   12103: 'Pump1: FeedPump: max. filling level drip pan', class Pump Warning Alarm, trigger "Pump1_FeedPump_DBW_2" bit 10
   12104: 'Pump1: FeedPump: dry-run protection', class Pump Warning Alarm, trigger "Pump1_FeedPump_DBW_2" bit 11
   12105: 'Pump1: FeedPump: incorrect time entry for runtime or pause time', class Pump Warning Alarm, trigger "Pump1_FeedPump_DBW_2" bit 12
   12106: 'Pump1: FeedPump: temperature for switch-off not reached', class Pump Warning Alarm, trigger "Pump1_FeedPump_DBW_2" bit 13
   12107: 'Pump1: FeedPump: fan motor protecting switch', class Pump Warning Alarm, trigger "Pump1_FeedPump_DBW_2" bit 14
   12108: 'Pump1: FeedPump: filling level too low', class Pump Warning Alarm, trigger "Pump1_FeedPump_DBW_2" bit 15
   12109: 'Pump1: FeedPump:', class Pump Warning Alarm, trigger "Pump1_FeedPump_DBW_2" bit 0
   12110: 'Pump1: FeedPump: filling selected but no barrel present', class Pump Warning Alarm, trigger "Pump1_FeedPump_DBW_2" bit 1
   12111: 'Pump1: FeedPump: no barrel present', class Pump Warning Alarm, trigger "Pump1_FeedPump_DBW_2" bit 2
   12112: 'Pump1: FeedPump:', class Pump Warning Alarm, trigger "Pump1_EdgeFilter_DBW_28" bit 8
   12113: 'Pump1: EdgeFilter: motor protecting switch has tripped', class Pump Warning Alarm, trigger "Pump1_EdgeFilter_DBW_28" bit 9
   12114: 'Pump1: EdgeFilter: max. differential pressure', class Pump Warning Alarm, trigger "Pump1_EdgeFilter_DBW_28" bit 10
   12115: 'Pump1: EdgeFilter: incorrect time entry for runtime or pause time', class Pump Warning Alarm, trigger "Pump1_EdgeFilter_DBW_28" bit 11
   12117: 'Pump1: Component pump: admission pressure not present', class Pump Archive Error Foaming, trigger "Pump1_Component_DBW_56" bit 8
   12118: 'Pump1: Component pump: motor protecting switch has tripped: Component pump', class Pump Error Alarm, trigger "Pump1_Component_DBW_56" bit 9
   12119: 'Pump1: Component pump: max. pressure', class Pump Archive Error Foaming, trigger "Pump1_Component_DBW_56" bit 10
   12120: 'Pump1: Component pump: pressure after feedpump too low', class Pump Error Alarm, trigger "Pump1_Component_DBW_56" bit 11
   12121: 'Pump1: Component pump: frequency converter fault', class Pump Error Alarm, trigger "Pump1_Component_DBW_56" bit 12
   12122: 'Pump1: Component pump: fan motor protecting switch', class Pump Warning Alarm, trigger "Pump1_Component_DBW_56" bit 13
   12123: 'Pump1: Component pump: min. tank filling level', class Pump Warning Alarm, trigger "Pump1_Component_DBW_56" bit 14
   12124: 'Pump1: Component pump: min. pressure not reached', class Pump Error Alarm, trigger "Pump1_Component_DBW_56" bit 15
   12125: 'Pump1: Component pump: pre-alarm, nitrogen', class Pump Warning Alarm, trigger "Pump1_Component_DBW_56" bit 0
   12126: 'Pump1: Component pump: flow- tolerance +', class Pump Warning Alarm, trigger "Pump1_Component_DBW_56" bit 1
   12127: 'Pump1: Component pump: flow tolerance -', class Pump Warning Alarm, trigger "Pump1_Component_DBW_56" bit 2
   12128: 'Pump1: Component pump: Timeout at fast pressure build-up', class Pump Warning Alarm, trigger "Pump1_Component_DBW_56" bit 3
   12129: 'Pump1: Component pump: enable temperature not reached', class Pump Warning Alarm, trigger "Pump1_Component_DBW_56" bit 4
   12130: 'Pump1: Component pump: converter restart delay active', class Pump Archive Warning Foaming, trigger "Pump1_Component_DBW_56" bit 5
   12131: 'Pump1: Component pump: alarm, nitrogen', class Pump Warning Alarm, trigger "Pump1_Component_DBW_56" bit 6
   12132: 'Pump1: Component pump: flow controller at limit', class Pump Warning Alarm, trigger "Pump1_Component_DBW_56" bit 7
   12133: 'Pump1: Component pump: component section was deselected', class Pump Warning Alarm, trigger "Pump1_Component_DBW_58" bit 8
   12134: 'Pump1: Component pump: deselected component section in interval', class Pump Warning Alarm, trigger "Pump1_Component_DBW_58" bit 9
   12135: 'Pump1: Component pump: fan motor protecting switch', class Pump Warning Alarm, trigger "Pump1_Component_DBW_58" bit 10
   12136: 'Pump1: Component pump: deselected component is required for entry', class Pump Warning Alarm, trigger "Pump1_Component_DBW_58" bit 11
   12137: 'Pump1: Component pump: flow controller at lower limit', class Pump Archive Warning Foaming, trigger "Pump1_Component_DBW_58" bit 12
   12138: 'Pump1: Component pump: max. filling level drip pan', class Pump Warning Alarm, trigger "Pump1_Component_DBW_58" bit 13
   12139: 'Pump1: Component pump:', class Pump Warning Alarm, trigger "Pump1_Component_DBW_58" bit 14
   12140: 'Pump1: Component pump:', class Pump Warning Alarm, trigger "Pump1_Component_DBW_58" bit 15
   12141: 'Pump1: Component pump:', class Pump Warning Alarm, trigger "Pump1_Component_DBW_58" bit 0
   12142: 'Pump1: Component pump:', class Pump Warning Alarm, trigger "Pump1_Component_DBW_58" bit 1
   12143: 'Pump1: Component pump:', class Pump Warning Alarm, trigger "Pump1_Component_DBW_58" bit 2
   12144: 'Pump1: Component pump:', class Pump Warning Alarm, trigger "Pump1_Component_DBW_58" bit 3
   12145: 'Pump1: Component pump:', class Pump Warning Alarm, trigger "Pump1_Component_DBW_58" bit 4
   12146: 'Pump1: Component pump:', class Pump Warning Alarm, trigger "Pump1_Component_DBW_58" bit 5
   12147: 'Pump1: Component pump:', class Pump Warning Alarm, trigger "Pump1_Component_DBW_58" bit 6
   12148: 'Pump1: Component pump:', class Pump Warning Alarm, trigger "Pump1_Component_DBW_58" bit 7
   12150: 'Pump1: Flow rate recording: measured value outside measuring range', class Pump Warning Alarm, trigger "Pump1_Flowrate_Record_DBW_106" bit 8
   12151: 'Pump1: Flow rate recording: warning, value exceeded', class Pump Warning Alarm, trigger "Pump1_Flowrate_Record_DBW_106" bit 9
   12152: 'Pump1: Flow rate recording: warning, value undershot', class Pump Warning Alarm, trigger "Pump1_Flowrate_Record_DBW_106" bit 10
   12153: 'Pump1: Flow rate recording: fault, value exceeded', class Pump Warning Alarm, trigger "Pump1_Flowrate_Record_DBW_106" bit 11
   12154: 'Pump1: Flow rate recording: fault, value undershot', class Pump Warning Alarm, trigger "Pump1_Flowrate_Record_DBW_106" bit 12
   12155: 'Pump1: Mixing ratio:', class Pump Warning Alarm, trigger "Pump1_Flowrate_Record_DBW_106" bit 0
   12156: 'Pump1: Mixing ratio: warning, value exceeded', class Pump Warning Alarm, trigger "Pump1_Flowrate_Record_DBW_106" bit 1
   12157: 'Pump1: Mixing ratio: warning, value undershot', class Pump Warning Alarm, trigger "Pump1_Flowrate_Record_DBW_106" bit 2
   12158: 'Pump1: Mixing ratio: fault, value exceeded', class Pump Error Alarm, trigger "Pump1_Flowrate_Record_DBW_106" bit 3
   12159: 'Pump1: Mixing ratio: fault, value undershot', class Pump Error Alarm, trigger "Pump1_Flowrate_Record_DBW_106" bit 4
   12160: 'Pump1: Pressure recording: measured value outside measuring range', class Pump Warning Alarm, trigger "Pump1_Pressure_Record_DBW_132" bit 8
   12161: 'Pump1: Pressure recording: warning, value exceeded', class Pump Warning Alarm, trigger "Pump1_Pressure_Record_DBW_132" bit 9
   12162: 'Pump1: Pressure recording: warning, value undershot', class Pump Warning Alarm, trigger "Pump1_Pressure_Record_DBW_132" bit 10
   12163: 'Pump1: Pressure recording: fault, value exceeded', class Pump Error Alarm, trigger "Pump1_Pressure_Record_DBW_132" bit 11
   12164: 'Pump1: Pressure recording: fault, value undershot', class Pump Error Alarm, trigger "Pump1_Pressure_Record_DBW_132" bit 12
   12165: 'Pump1: Temp. recording HP heat exch.: measured value outside measuring range', class Pump Warning Alarm, trigger "Pump1_Heatexchanger_DBW_210" bit 8
   12166: 'Pump1: Temp. recording HP heat exch.: warning, value exceeded', class Pump Warning Alarm, trigger "Pump1_Heatexchanger_DBW_210" bit 9
   12167: 'Pump1: Temp. recording HP heat exch.: warning, value undershot', class Pump Warning Alarm, trigger "Pump1_Heatexchanger_DBW_210" bit 10
   12168: 'Pump1: Temp. recording HP heat exch.: fault, value exceeded', class Pump Error Alarm, trigger "Pump1_Heatexchanger_DBW_210" bit 11
   12169: 'Pump1: Temp. recording HP heat exch.: fault, value undershot', class Pump Error Alarm, trigger "Pump1_Heatexchanger_DBW_210" bit 12
   12201: 'Pump2: FeedPump: motor protecting switch has tripped', class Pump Warning Alarm, trigger "Pump2_FeedPump_DBW_4" bit 8
   12202: 'Pump2: FeedPump: frequency converter fault', class Pump Warning Alarm, trigger "Pump2_FeedPump_DBW_4" bit 9
   12203: 'Pump2: FeedPump: max. filling level drip pan', class Pump Warning Alarm, trigger "Pump2_FeedPump_DBW_4" bit 10
   12204: 'Pump2: FeedPump: dry-run protection', class Pump Warning Alarm, trigger "Pump2_FeedPump_DBW_4" bit 11
   12205: 'Pump2: FeedPump: incorrect time entry for runtime or pause time', class Pump Warning Alarm, trigger "Pump2_FeedPump_DBW_4" bit 12
   12206: 'Pump2: FeedPump: temperature for switch-off not reached', class Pump Warning Alarm, trigger "Pump2_FeedPump_DBW_4" bit 13
   12207: 'Pump2: FeedPump: fan motor protecting switch', class Pump Warning Alarm, trigger "Pump2_FeedPump_DBW_4" bit 14
   12208: 'Pump2: FeedPump: filling level too low', class Pump Warning Alarm, trigger "Pump2_FeedPump_DBW_4" bit 15
   12209: 'Pump2: FeedPump:', class Pump Warning Alarm, trigger "Pump2_FeedPump_DBW_4" bit 0
   12210: 'Pump2: FeedPump: filling selected but no barrel present', class Pump Warning Alarm, trigger "Pump2_FeedPump_DBW_4" bit 1
   12211: 'Pump2: FeedPump: no barrel present', class Pump Warning Alarm, trigger "Pump2_FeedPump_DBW_4" bit 2
   12212: 'Pump2: FeedPump:', class Pump Warning Alarm, trigger "Pump2_FeedPump_DBW_4" bit 3
   12213: 'Pump2: EdgeFilter: motor protecting switch has tripped', class Pump Warning Alarm, trigger "Pump2_EdgeFilter_DBW_30" bit 8
   12214: 'Pump2: EdgeFilter: max. differential pressure', class Pump Warning Alarm, trigger "Pump2_EdgeFilter_DBW_30" bit 9
   12215: 'Pump2: EdgeFilter: incorrect time entry for runtime or pause time', class Pump Warning Alarm, trigger "Pump2_EdgeFilter_DBW_30" bit 10
   12216: 'Pump2: EdgeFilter:', class Pump Warning Alarm, trigger "Pump2_EdgeFilter_DBW_30" bit 11
   12217: 'Pump2: Component pump: admission pressure not present', class Pump Archive Error Foaming, trigger "Pump2_Component_DBW_60" bit 8
   12218: 'Pump2: Component pump: motor protecting switch has tripped: Component pump', class Pump Error Alarm, trigger "Pump2_Component_DBW_60" bit 9
   12219: 'Pump2: Component pump: max. pressure', class Pump Error Alarm, trigger "Pump2_Component_DBW_60" bit 10
   12220: 'Pump2: Component pump: pressure after feedpump too low', class Pump Error Alarm, trigger "Pump2_Component_DBW_60" bit 11
   12221: 'Pump2: Component pump: frequency converter fault', class Pump Archive Warning Foaming, trigger "Pump2_Component_DBW_60" bit 12
   12222: 'Pump2: Component pump: fan motor protecting switch', class Pump Warning Alarm, trigger "Pump2_Component_DBW_60" bit 13
   12223: 'Pump2: Component pump: min. tank filling level', class Pump Warning Alarm, trigger "Pump2_Component_DBW_60" bit 14
   12224: 'Pump2: Component pump: min. pressure not reached', class Pump Archive Error Foaming, trigger "Pump2_Component_DBW_60" bit 15
   12225: 'Pump2: Component pump: pre-alarm, nitrogen', class Pump Warning Alarm, trigger "Pump2_Component_DBW_60" bit 0
   12226: 'Pump2: Component pump: flow- tolerance +', class Pump Warning Alarm, trigger "Pump2_Component_DBW_60" bit 1
   12227: 'Pump2: Component pump: flow tolerance -', class Pump Warning Alarm, trigger "Pump2_Component_DBW_60" bit 2
   12228: 'Pump2: Component pump: Timeout at fast pressure build-up', class Pump Warning Alarm, trigger "Pump2_Component_DBW_60" bit 3
   12229: 'Pump2: Component pump: enable temperature not reached', class Pump Warning Alarm, trigger "Pump2_Component_DBW_60" bit 4
   12230: 'Pump2: Component pump: converter restart delay active', class Pump Archive Warning Foaming, trigger "Pump2_Component_DBW_60" bit 5
   12231: 'Pump2: Component pump: alarm, nitrogen', class Pump Warning Alarm, trigger "Pump2_Component_DBW_60" bit 6
   12232: 'Pump2: Component pump: flow controller at limit', class Pump Warning Alarm, trigger "Pump2_Component_DBW_60" bit 7
   12233: 'Pump2: Component pump: component section was deselected', class Pump Warning Alarm, trigger "Pump2_Component_DBW_62" bit 8
   12234: 'Pump2: Component pump: deselected component section in interval', class Pump Warning Alarm, trigger "Pump2_Component_DBW_62" bit 9
   12235: 'Pump2: Component pump: fan motor protecting switch', class Pump Warning Alarm, trigger "Pump2_Component_DBW_62" bit 10
   12236: 'Pump2: Component pump: deselected component is required for entry', class Pump Warning Alarm, trigger "Pump2_Component_DBW_62" bit 11
   12237: 'Pump2: Component pump: flow controller at lower limit', class Pump Archive Warning Foaming, trigger "Pump2_Component_DBW_62" bit 12
   12238: 'Pump2: Component pump: max. filling level drip pan', class Pump Warning Alarm, trigger "Pump2_Component_DBW_62" bit 13
   12239: 'Pump2: Component pump:', class Pump Warning Alarm, trigger "Pump2_Component_DBW_62" bit 14
   12240: 'Pump2: Component pump:', class Pump Warning Alarm, trigger "Pump2_Component_DBW_62" bit 15
   12241: 'Pump2: Component pump:', class Pump Warning Alarm, trigger "Pump2_Component_DBW_62" bit 0
   12242: 'Pump2: Component pump:', class Pump Warning Alarm, trigger "Pump2_Component_DBW_62" bit 1
   12243: 'Pump2: Component pump:', class Pump Warning Alarm, trigger "Pump2_Component_DBW_62" bit 2
   12244: 'Pump2: Component pump:', class Pump Warning Alarm, trigger "Pump2_Component_DBW_62" bit 3
   12245: 'Pump2: Component pump:', class Pump Warning Alarm, trigger "Pump2_Component_DBW_62" bit 4
   12246: 'Pump2: Component pump:', class Pump Warning Alarm, trigger "Pump2_Component_DBW_62" bit 5
   12247: 'Pump2: Component pump:', class Pump Warning Alarm, trigger "Pump2_Component_DBW_62" bit 6
   12248: 'Pump2: Component pump:', class Pump Warning Alarm, trigger "Pump2_Component_DBW_62" bit 7
   12116: 'Pump1: EdgeFilter:', class Pump Warning Alarm, trigger "Pump1_EdgeFilter_DBW_28" bit 12
   12250: 'Pump2: Flow rate recording: measured value outside measuring range', class Pump Warning Alarm, trigger "Pump2_Flowrate_Record_DBW_108" bit 8
   12251: 'Pump2: Flow rate recording: warning, value exceeded', class Pump Warning Alarm, trigger "Pump2_Flowrate_Record_DBW_108" bit 9
   12252: 'Pump2: Flow rate recording: warning, value undershot', class Pump Warning Alarm, trigger "Pump2_Flowrate_Record_DBW_108" bit 10
   12253: 'Pump2: Flow rate recording: fault, value exceeded', class Pump Error Alarm, trigger "Pump2_Flowrate_Record_DBW_108" bit 11
   12254: 'Pump2: Flow rate recording: fault, value undershot', class Pump Error Alarm, trigger "Pump2_Flowrate_Record_DBW_108" bit 12
   12255: 'Pump2: Mixing ratio:', class Pump Warning Alarm, trigger "Pump2_Flowrate_Record_DBW_108" bit 0
   12256: 'Pump2: Mixing ratio: warning, value exceeded', class Pump Warning Alarm, trigger "Pump2_Flowrate_Record_DBW_108" bit 1
   12257: 'Pump2: Mixing ratio: warning, value undershot', class Pump Warning Alarm, trigger "Pump2_Flowrate_Record_DBW_108" bit 2
   12258: 'Pump2: Mixing ratio: fault, value exceeded', class Pump Error Alarm, trigger "Pump2_Flowrate_Record_DBW_108" bit 3
   12259: 'Pump2: Mixing ratio: fault, value undershot', class Pump Error Alarm, trigger "Pump2_Flowrate_Record_DBW_108" bit 4
   12260: 'Pump2: Pressure recording: measured value outside measuring range', class Pump Warning Alarm, trigger "Pump2_Pressure_Record_DBW_134" bit 8
   12261: 'Pump2: Pressure recording: warning, value exceeded', class Pump Warning Alarm, trigger "Pump2_Pressure_Record_DBW_134" bit 9
   12262: 'Pump2: Pressure recording: warning, value undershot', class Pump Warning Alarm, trigger "Pump2_Pressure_Record_DBW_134" bit 10
   12263: 'Pump2: Pressure recording: fault, value exceeded', class Pump Error Alarm, trigger "Pump2_Pressure_Record_DBW_134" bit 11
   12264: 'Pump2: Pressure recording: fault, value undershot', class Pump Error Alarm, trigger "Pump2_Pressure_Record_DBW_134" bit 12
   12265: 'Pump2: Temp. recording HP heat exch.: measured value outside measuring range', class Pump Warning Alarm, trigger "Pump2_Heatexchanger_DBW_212" bit 8
   12266: 'Pump2: Temp. recording HP heat exch.: warning, value exceeded', class Pump Warning Alarm, trigger "Pump2_Heatexchanger_DBW_212" bit 9
   12267: 'Pump2: Temp. recording HP heat exch.: warning, value undershot', class Pump Warning Alarm, trigger "Pump2_Heatexchanger_DBW_212" bit 10
   12268: 'Pump2: Temp. recording HP heat exch.: fault, value exceeded', class Pump Error Alarm, trigger "Pump2_Heatexchanger_DBW_212" bit 11
   12269: 'Pump2: Temp. recording HP heat exch.: fault, value undershot', class Pump Error Alarm, trigger "Pump2_Heatexchanger_DBW_212" bit 12
   12301: 'Pump3: FeedPump: motor protecting switch has tripped', class Pump Warning Alarm, trigger "Pump3_FeedPump_DBW_6" bit 8
   12302: 'Pump3: FeedPump: frequency converter fault', class Pump Warning Alarm, trigger "Pump3_FeedPump_DBW_6" bit 9
   12303: 'Pump3: FeedPump: max. filling level drip pan', class Pump Warning Alarm, trigger "Pump3_FeedPump_DBW_6" bit 10
   12304: 'Pump3: FeedPump: dry-run protection', class Pump Warning Alarm, trigger "Pump3_FeedPump_DBW_6" bit 11
   12305: 'Pump3: FeedPump: incorrect time entry for runtime or pause time', class Pump Warning Alarm, trigger "Pump3_FeedPump_DBW_6" bit 12
   12306: 'Pump3: FeedPump: temperature for switch-off not reached', class Pump Warning Alarm, trigger "Pump3_FeedPump_DBW_6" bit 13
   12307: 'Pump3: FeedPump: fan motor protecting switch', class Pump Warning Alarm, trigger "Pump3_FeedPump_DBW_6" bit 14
   12308: 'Pump3: FeedPump: filling level too low', class Pump Warning Alarm, trigger "Pump3_FeedPump_DBW_6" bit 15
   12309: 'Pump3: FeedPump:', class Pump Warning Alarm, trigger "Pump3_FeedPump_DBW_6" bit 0
   12310: 'Pump3: FeedPump: filling selected but no barrel present', class Pump Warning Alarm, trigger "Pump3_FeedPump_DBW_6" bit 1
   12311: 'Pump3: FeedPump: no barrel present', class Pump Warning Alarm, trigger "Pump3_FeedPump_DBW_6" bit 2
   12312: 'Pump3: FeedPump:', class Pump Warning Alarm, trigger "Pump3_FeedPump_DBW_6" bit 3
   12313: 'Pump3: EdgeFilter: motor protecting switch has tripped', class Pump Warning Alarm, trigger "Pump3_EdgeFilter_DBW_32" bit 8
   12314: 'Pump3: EdgeFilter: max. differential pressure', class Pump Warning Alarm, trigger "Pump3_EdgeFilter_DBW_32" bit 9
   12315: 'Pump3: EdgeFilter: incorrect time entry for runtime or pause time', class Pump Warning Alarm, trigger "Pump3_EdgeFilter_DBW_32" bit 10
   12316: 'Pump3: EdgeFilter:', class Pump Warning Alarm, trigger "Pump3_EdgeFilter_DBW_32" bit 11
   12317: 'Pump3: Component pump: admission pressure not present', class Pump Error Alarm, trigger "Pump3_Component_DBW_64" bit 8
   12318: 'Pump3: Component pump: motor protecting switch has tripped: Component pump', class Pump Error Alarm, trigger "Pump3_Component_DBW_64" bit 9
   12319: 'Pump3: Component pump: max. pressure', class Pump Error Alarm, trigger "Pump3_Component_DBW_64" bit 10
   12320: 'Pump3: Component pump: pressure after feedpump too low', class Pump Error Alarm, trigger "Pump3_Component_DBW_64" bit 11
   12321: 'Pump3: Component pump: frequency converter fault', class Pump Warning Alarm, trigger "Pump3_Component_DBW_64" bit 12
   12322: 'Pump3: Component pump: fan motor protecting switch', class Pump Warning Alarm, trigger "Pump3_Component_DBW_64" bit 13
   12323: 'Pump3: Component pump: min. tank filling level', class Pump Warning Alarm, trigger "Pump3_Component_DBW_64" bit 14
   12324: 'Pump3: Component pump: min. pressure not reached', class Pump Error Alarm, trigger "Pump3_Component_DBW_64" bit 15
   12325: 'Pump3: Component pump: pre-alarm, nitrogen', class Pump Warning Alarm, trigger "Pump3_Component_DBW_64" bit 0
   12326: 'Pump3: Component pump: flow- tolerance +', class Pump Warning Alarm, trigger "Pump3_Component_DBW_64" bit 1
   12327: 'Pump3: Component pump: flow tolerance -', class Pump Warning Alarm, trigger "Pump3_Component_DBW_64" bit 2
   12328: 'Pump3: Component pump: Timeout at fast pressure build-up', class Pump Warning Alarm, trigger "Pump3_Component_DBW_64" bit 3
   12329: 'Pump3: Component pump: enable temperature not reached', class Pump Warning Alarm, trigger "Pump3_Component_DBW_64" bit 4
   12330: 'Pump3: Component pump: converter restart delay active', class Pump Warning Alarm, trigger "Pump3_Component_DBW_64" bit 5
   12331: 'Pump3: Component pump: alarm, nitrogen', class Pump Warning Alarm, trigger "Pump3_Component_DBW_64" bit 6
   12332: 'Pump3: Component pump: flow controller at limit', class Pump Warning Alarm, trigger "Pump3_Component_DBW_64" bit 7
   12333: 'Pump3: Component pump: component section was deselected', class Pump Warning Alarm, trigger "Pump3_Component_DBW_66" bit 8
   12334: 'Pump3: Component pump: deselected component section in interval', class Pump Warning Alarm, trigger "Pump3_Component_DBW_66" bit 9
   12335: 'Pump3: Component pump: fan motor protecting switch', class Pump Warning Alarm, trigger "Pump3_Component_DBW_66" bit 10
   12336: 'Pump3: Component pump: deselected component is required for entry', class Pump Warning Alarm, trigger "Pump3_Component_DBW_66" bit 11
   12337: 'Pump3: Component pump: flow controller at lower limit', class Pump Warning Alarm, trigger "Pump3_Component_DBW_66" bit 12
   12338: 'Pump3: Component pump: max. filling level drip pan', class Pump Warning Alarm, trigger "Pump3_Component_DBW_66" bit 13
   12339: 'Pump3: Component pump:', class Pump Warning Alarm, trigger "Pump3_Component_DBW_66" bit 14
   12340: 'Pump3: Component pump:', class Pump Warning Alarm, trigger "Pump3_Component_DBW_66" bit 15
   12341: 'Pump3: Component pump:', class Pump Warning Alarm, trigger "Pump3_Component_DBW_66" bit 0
   12342: 'Pump3: Component pump:', class Pump Warning Alarm, trigger "Pump3_Component_DBW_66" bit 1
   12343: 'Pump3: Component pump:', class Pump Warning Alarm, trigger "Pump3_Component_DBW_66" bit 2
   12344: 'Pump3: Component pump:', class Pump Warning Alarm, trigger "Pump3_Component_DBW_66" bit 3
   12345: 'Pump3: Component pump:', class Pump Warning Alarm, trigger "Pump3_Component_DBW_66" bit 4
   12346: 'Pump3: Component pump:', class Pump Warning Alarm, trigger "Pump3_Component_DBW_66" bit 5
   12347: 'Pump3: Component pump:', class Pump Warning Alarm, trigger "Pump3_Component_DBW_66" bit 6
   12348: 'Pump3: Component pump:', class Pump Warning Alarm, trigger "Pump3_Component_DBW_66" bit 7
   12350: 'Pump3: Flow rate recording: measured value outside measuring range', class Pump Warning Alarm, trigger "Pump3_Flowrate_Record_DBW_110" bit 8
   12351: 'Pump3: Flow rate recording: warning, value exceeded', class Pump Warning Alarm, trigger "Pump3_Flowrate_Record_DBW_110" bit 9
   12352: 'Pump3: Flow rate recording: warning, value undershot', class Pump Warning Alarm, trigger "Pump3_Flowrate_Record_DBW_110" bit 10
   12353: 'Pump3: Flow rate recording: fault, value exceeded', class Pump Error Alarm, trigger "Pump3_Flowrate_Record_DBW_110" bit 11
   12354: 'Pump3: Flow rate recording: fault, value undershot', class Pump Error Alarm, trigger "Pump3_Flowrate_Record_DBW_110" bit 12
   12355: 'Pump3: Mixing ratio:', class Pump Warning Alarm, trigger "Pump3_Flowrate_Record_DBW_110" bit 0
   12356: 'Pump3: Mixing ratio: warning, value exceeded', class Pump Warning Alarm, trigger "Pump3_Flowrate_Record_DBW_110" bit 1
   12357: 'Pump3: Mixing ratio: warning, value undershot', class Pump Warning Alarm, trigger "Pump3_Flowrate_Record_DBW_110" bit 2
   12358: 'Pump3: Mixing ratio: fault, value exceeded', class Pump Error Alarm, trigger "Pump3_Flowrate_Record_DBW_110" bit 3
   12359: 'Pump3: Mixing ratio: fault, value undershot', class Pump Error Alarm, trigger "Pump3_Flowrate_Record_DBW_110" bit 4
   12360: 'Pump3: Pressure recording: measured value outside measuring range', class Pump Warning Alarm, trigger "Pump3_Pressure_Record_DBW_136" bit 8
   12361: 'Pump3: Pressure recording: warning, value exceeded', class Pump Warning Alarm, trigger "Pump3_Pressure_Record_DBW_136" bit 9
   12362: 'Pump3: Pressure recording: warning, value undershot', class Pump Warning Alarm, trigger "Pump3_Pressure_Record_DBW_136" bit 10
   12363: 'Pump3: Pressure recording: fault, value exceeded', class Pump Error Alarm, trigger "Pump3_Pressure_Record_DBW_136" bit 11
   12364: 'Pump3: Pressure recording: fault, value undershot', class Pump Error Alarm, trigger "Pump3_Pressure_Record_DBW_136" bit 12
   12365: 'Pump3: Temp. recording HP heat exch.: measured value outside measuring range', class Pump Warning Alarm, trigger "Pump3_Heatexchanger_DBW_214" bit 8
   12366: 'Pump3: Temp. recording HP heat exch.: warning, value exceeded', class Pump Warning Alarm, trigger "Pump3_Heatexchanger_DBW_214" bit 9
   12367: 'Pump3: Temp. recording HP heat exch.: warning, value undershot', class Pump Warning Alarm, trigger "Pump3_Heatexchanger_DBW_214" bit 10
   12368: 'Pump3: Temp. recording HP heat exch.: fault, value exceeded', class Pump Error Alarm, trigger "Pump3_Heatexchanger_DBW_214" bit 11
   12369: 'Pump3: Temp. recording HP heat exch.: fault, value undershot', class Pump Error Alarm, trigger "Pump3_Heatexchanger_DBW_214" bit 12
   12401: 'Pump4: FeedPump: motor protecting switch has tripped', class Pump Warning Alarm, trigger "Pump4_FeedPump_DBW_8" bit 8
   12402: 'Pump4: FeedPump: frequency converter fault', class Pump Warning Alarm, trigger "Pump4_FeedPump_DBW_8" bit 9
   12403: 'Pump4: FeedPump: max. filling level drip pan', class Pump Warning Alarm, trigger "Pump4_FeedPump_DBW_8" bit 10
   12404: 'Pump4: FeedPump: dry-run protection', class Pump Warning Alarm, trigger "Pump4_FeedPump_DBW_8" bit 11
   12405: 'Pump4: FeedPump: incorrect time entry for runtime or pause time', class Pump Warning Alarm, trigger "Pump4_FeedPump_DBW_8" bit 12
   12406: 'Pump4: FeedPump: temperature for switch-off not reached', class Pump Warning Alarm, trigger "Pump4_FeedPump_DBW_8" bit 13
   12407: 'Pump4: FeedPump: fan motor protecting switch', class Pump Warning Alarm, trigger "Pump4_FeedPump_DBW_8" bit 14
   12408: 'Pump4: FeedPump: filling level too low', class Pump Warning Alarm, trigger "Pump4_FeedPump_DBW_8" bit 15
   12409: 'Pump4: FeedPump:', class Pump Warning Alarm, trigger "Pump4_FeedPump_DBW_8" bit 0
   12410: 'Pump4: FeedPump: filling selected but no barrel present', class Pump Warning Alarm, trigger "Pump4_FeedPump_DBW_8" bit 1
   12411: 'Pump4: FeedPump: no barrel present', class Pump Warning Alarm, trigger "Pump4_FeedPump_DBW_8" bit 2
   12412: 'Pump4: FeedPump:', class Pump Warning Alarm, trigger "Pump4_FeedPump_DBW_8" bit 3
   12413: 'Pump4: EdgeFilter: motor protecting switch has tripped', class Pump Warning Alarm, trigger "Pump4_EdgeFilter_DBW_34" bit 8
   12414: 'Pump4: EdgeFilter: max. differential pressure', class Pump Warning Alarm, trigger "Pump4_EdgeFilter_DBW_34" bit 9
   12415: 'Pump4: EdgeFilter: incorrect time entry for runtime or pause time', class Pump Warning Alarm, trigger "Pump4_EdgeFilter_DBW_34" bit 10
   12416: 'Pump4: EdgeFilter:', class Pump Warning Alarm, trigger "Pump4_EdgeFilter_DBW_34" bit 11
   12417: 'Pump4: Component pump: admission pressure not present', class Pump Error Alarm, trigger "Pump4_Component_DBW_68" bit 8
   12418: 'Pump4: Component pump: motor protecting switch has tripped: Component pump', class Pump Error Alarm, trigger "Pump4_Component_DBW_68" bit 9
   12419: 'Pump4: Component pump: max. pressure', class Pump Error Alarm, trigger "Pump4_Component_DBW_68" bit 10
   12420: 'Pump4: Component pump: pressure after feedpump too low', class Pump Error Alarm, trigger "Pump4_Component_DBW_68" bit 11
   12421: 'Pump4: Component pump: frequency converter fault', class Pump Warning Alarm, trigger "Pump4_Component_DBW_68" bit 12
   12422: 'Pump4: Component pump: fan motor protecting switch', class Pump Warning Alarm, trigger "Pump4_Component_DBW_68" bit 13
   12423: 'Pump4: Component pump: min. tank filling level', class Pump Warning Alarm, trigger "Pump4_Component_DBW_68" bit 14
   12424: 'Pump4: Component pump: min. pressure not reached', class Pump Error Alarm, trigger "Pump4_Component_DBW_68" bit 15
   12425: 'Pump4: Component pump: pre-alarm, nitrogen', class Pump Warning Alarm, trigger "Pump4_Component_DBW_68" bit 0
   12426: 'Pump4: Component pump: flow- tolerance +', class Pump Warning Alarm, trigger "Pump4_Component_DBW_68" bit 1
   12427: 'Pump4: Component pump: flow tolerance -', class Pump Warning Alarm, trigger "Pump4_Component_DBW_68" bit 2
   12428: 'Pump4: Component pump: Timeout at fast pressure build-up', class Pump Warning Alarm, trigger "Pump4_Component_DBW_68" bit 3
   12429: 'Pump4: Component pump: enable temperature not reached', class Pump Warning Alarm, trigger "Pump4_Component_DBW_68" bit 4
   12430: 'Pump4: Component pump: converter restart delay active', class Pump Warning Alarm, trigger "Pump4_Component_DBW_68" bit 5
   12431: 'Pump4: Component pump: alarm, nitrogen', class Pump Warning Alarm, trigger "Pump4_Component_DBW_68" bit 6
   12432: 'Pump4: Component pump: flow controller at limit', class Pump Warning Alarm, trigger "Pump4_Component_DBW_68" bit 7
   12433: 'Pump4: Component pump: component section was deselected', class Pump Warning Alarm, trigger "Pump4_Component_DBW_70" bit 8
   12434: 'Pump4: Component pump: deselected component section in interval', class Pump Warning Alarm, trigger "Pump4_Component_DBW_70" bit 9
   12435: 'Pump4: Component pump: fan motor protecting switch', class Pump Warning Alarm, trigger "Pump4_Component_DBW_70" bit 10
   12436: 'Pump4: Component pump: deselected component is required for entry', class Pump Warning Alarm, trigger "Pump4_Component_DBW_70" bit 11
   12437: 'Pump4: Component pump: flow controller at lower limit', class Pump Warning Alarm, trigger "Pump4_Component_DBW_70" bit 12
   12438: 'Pump4: Component pump: max. filling level drip pan', class Pump Warning Alarm, trigger "Pump4_Component_DBW_70" bit 13
   12439: 'Pump4: Component pump:', class Pump Warning Alarm, trigger "Pump4_Component_DBW_70" bit 14
   12440: 'Pump4: Component pump:', class Pump Warning Alarm, trigger "Pump4_Component_DBW_70" bit 15
   12441: 'Pump4: Component pump:', class Pump Warning Alarm, trigger "Pump4_Component_DBW_70" bit 0
   12442: 'Pump4: Component pump:', class Pump Warning Alarm, trigger "Pump4_Component_DBW_70" bit 1
   12443: 'Pump4: Component pump:', class Pump Warning Alarm, trigger "Pump4_Component_DBW_70" bit 2
   12444: 'Pump4: Component pump:', class Pump Warning Alarm, trigger "Pump4_Component_DBW_70" bit 3
   12445: 'Pump4: Component pump:', class Pump Warning Alarm, trigger "Pump4_Component_DBW_70" bit 4
   12446: 'Pump4: Component pump:', class Pump Warning Alarm, trigger "Pump4_Component_DBW_70" bit 5
   12447: 'Pump4: Component pump:', class Pump Warning Alarm, trigger "Pump4_Component_DBW_70" bit 6
   12448: 'Pump4: Component pump:', class Pump Warning Alarm, trigger "Pump4_Component_DBW_70" bit 7
   12450: 'Pump4: Flow rate recording: measured value outside measuring range', class Pump Warning Alarm, trigger "Pump4_Flowrate_Record_DBW_112" bit 8
   12451: 'Pump4: Flow rate recording: warning, value exceeded', class Pump Warning Alarm, trigger "Pump4_Flowrate_Record_DBW_112" bit 9
   12452: 'Pump4: Flow rate recording: warning, value undershot', class Pump Warning Alarm, trigger "Pump4_Flowrate_Record_DBW_112" bit 10
   12453: 'Pump4: Flow rate recording: fault, value exceeded', class Pump Error Alarm, trigger "Pump4_Flowrate_Record_DBW_112" bit 11
   12454: 'Pump4: Flow rate recording: fault, value undershot', class Pump Error Alarm, trigger "Pump4_Flowrate_Record_DBW_112" bit 12
   12455: 'Pump4: Mixing ratio:', class Pump Warning Alarm, trigger "Pump4_Flowrate_Record_DBW_112" bit 0
   12456: 'Pump4: Mixing ratio: warning, value exceeded', class Pump Warning Alarm, trigger "Pump4_Flowrate_Record_DBW_112" bit 1
   12457: 'Pump4: Mixing ratio: warning, value undershot', class Pump Warning Alarm, trigger "Pump4_Flowrate_Record_DBW_112" bit 2
   12458: 'Pump4: Mixing ratio: fault, value exceeded', class Pump Error Alarm, trigger "Pump4_Flowrate_Record_DBW_112" bit 3
   12459: 'Pump4: Mixing ratio: fault, value undershot', class Pump Error Alarm, trigger "Pump4_Flowrate_Record_DBW_112" bit 4
   12460: 'Pump4: Pressure recording: measured value outside measuring range', class Pump Warning Alarm, trigger "Pump4_Pressure_Record_DBW_138" bit 8
   12461: 'Pump4: Pressure recording: warning, value exceeded', class Pump Warning Alarm, trigger "Pump4_Pressure_Record_DBW_138" bit 9
   12462: 'Pump4: Pressure recording: warning, value undershot', class Pump Warning Alarm, trigger "Pump4_Pressure_Record_DBW_138" bit 10
   12463: 'Pump4: Pressure recording: fault, value exceeded', class Pump Error Alarm, trigger "Pump4_Pressure_Record_DBW_138" bit 11
   12464: 'Pump4: Pressure recording: fault, value undershot', class Pump Error Alarm, trigger "Pump4_Pressure_Record_DBW_138" bit 12
   12465: 'Pump4: Temp. recording HP heat exch.: measured value outside measuring range', class Pump Warning Alarm, trigger "Pump4_Heatexchanger_DBW_216" bit 8
   12466: 'Pump4: Temp. recording HP heat exch.: warning, value exceeded', class Pump Warning Alarm, trigger "Pump4_Heatexchanger_DBW_216" bit 9
   12467: 'Pump4: Temp. recording HP heat exch.: warning, value undershot', class Pump Warning Alarm, trigger "Pump4_Heatexchanger_DBW_216" bit 10
   12468: 'Pump4: Temp. recording HP heat exch.: fault, value exceeded', class Pump Error Alarm, trigger "Pump4_Heatexchanger_DBW_216" bit 11
   12469: 'Pump4: Temp. recording HP heat exch.: fault, value undershot', class Pump Error Alarm, trigger "Pump4_Heatexchanger_DBW_216" bit 12
   12501: 'Pump5: FeedPump: motor protecting switch has tripped', class Pump Warning Alarm, trigger "Pump5_FeedPump_DBW_10" bit 8
   12502: 'Pump5: FeedPump: frequency converter fault', class Pump Warning Alarm, trigger "Pump5_FeedPump_DBW_10" bit 9
   12503: 'Pump5: FeedPump: max. filling level drip pan', class Pump Warning Alarm, trigger "Pump5_FeedPump_DBW_10" bit 10
   12504: 'Pump5: FeedPump: dry-run protection', class Pump Warning Alarm, trigger "Pump5_FeedPump_DBW_10" bit 11
   12505: 'Pump5: FeedPump: incorrect time entry for runtime or pause time', class Pump Warning Alarm, trigger "Pump5_FeedPump_DBW_10" bit 12
   12506: 'Pump5: FeedPump: temperature for switch-off not reached', class Pump Warning Alarm, trigger "Pump5_FeedPump_DBW_10" bit 13
   12507: 'Pump5: FeedPump: fan motor protecting switch', class Pump Warning Alarm, trigger "Pump5_FeedPump_DBW_10" bit 14
   12508: 'Pump5: FeedPump: filling level too low', class Pump Warning Alarm, trigger "Pump5_FeedPump_DBW_10" bit 15
   12509: 'Pump5: FeedPump:', class Pump Warning Alarm, trigger "Pump5_FeedPump_DBW_10" bit 0
   12510: 'Pump5: FeedPump: filling selected but no barrel present', class Pump Warning Alarm, trigger "Pump5_FeedPump_DBW_10" bit 1
   12511: 'Pump5: FeedPump: no barrel present', class Pump Warning Alarm, trigger "Pump5_FeedPump_DBW_10" bit 2
   12512: 'Pump5: FeedPump:', class Pump Warning Alarm, trigger "Pump5_FeedPump_DBW_10" bit 3
   12513: 'Pump5: EdgeFilter: motor protecting switch has tripped', class Pump Warning Alarm, trigger "Pump5_EdgeFilter_DBW_36" bit 8
   12514: 'Pump5: EdgeFilter: max. differential pressure', class Pump Warning Alarm, trigger "Pump5_EdgeFilter_DBW_36" bit 9
   12515: 'Pump5: EdgeFilter: incorrect time entry for runtime or pause time', class Pump Warning Alarm, trigger "Pump5_EdgeFilter_DBW_36" bit 10
   12516: 'Pump5: EdgeFilter:', class Pump Warning Alarm, trigger "Pump5_EdgeFilter_DBW_36" bit 11
   12517: 'Pump5: Component pump: admission pressure not present', class Pump Error Alarm, trigger "Pump5_Component_DBW_72" bit 8
   12518: 'Pump5: Component pump: motor protecting switch has tripped: Component pump', class Pump Error Alarm, trigger "Pump5_Component_DBW_72" bit 9
   12519: 'Pump5: Component pump: max. pressure', class Pump Error Alarm, trigger "Pump5_Component_DBW_72" bit 10
   12520: 'Pump5: Component pump: pressure after feedpump too low', class Pump Error Alarm, trigger "Pump5_Component_DBW_72" bit 11
   12521: 'Pump5: Component pump: frequency converter fault', class Pump Warning Alarm, trigger "Pump5_Component_DBW_72" bit 12
   12522: 'Pump5: Component pump: fan motor protecting switch', class Pump Warning Alarm, trigger "Pump5_Component_DBW_72" bit 13
   12523: 'Pump5: Component pump: min. tank filling level', class Pump Warning Alarm, trigger "Pump5_Component_DBW_72" bit 14
   12524: 'Pump5: Component pump: min. pressure not reached', class Pump Error Alarm, trigger "Pump5_Component_DBW_72" bit 15
   12525: 'Pump5: Component pump: pre-alarm, nitrogen', class Pump Warning Alarm, trigger "Pump5_Component_DBW_72" bit 0
   12526: 'Pump5: Component pump: flow- tolerance +', class Pump Warning Alarm, trigger "Pump5_Component_DBW_72" bit 1
   12527: 'Pump5: Component pump: flow tolerance -', class Pump Warning Alarm, trigger "Pump5_Component_DBW_72" bit 2
   12528: 'Pump5: Component pump: Timeout at fast pressure build-up', class Pump Warning Alarm, trigger "Pump5_Component_DBW_72" bit 3
   12529: 'Pump5: Component pump: enable temperature not reached', class Pump Warning Alarm, trigger "Pump5_Component_DBW_72" bit 4
   12530: 'Pump5: Component pump: converter restart delay active', class Pump Warning Alarm, trigger "Pump5_Component_DBW_72" bit 5
   12531: 'Pump5: Component pump: alarm, nitrogen', class Pump Warning Alarm, trigger "Pump5_Component_DBW_72" bit 6
   12532: 'Pump5: Component pump: flow controller at limit', class Pump Warning Alarm, trigger "Pump5_Component_DBW_72" bit 7
   12533: 'Pump5: Component pump: component section was deselected', class Pump Warning Alarm, trigger "Pump5_Component_DBW_74" bit 8
   12534: 'Pump5: Component pump: deselected component section in interval', class Pump Warning Alarm, trigger "Pump5_Component_DBW_74" bit 9
   12535: 'Pump5: Component pump: fan motor protecting switch', class Pump Warning Alarm, trigger "Pump5_Component_DBW_74" bit 10
   12536: 'Pump5: Component pump: deselected component is required for entry', class Pump Warning Alarm, trigger "Pump5_Component_DBW_74" bit 11
   12537: 'Pump5: Component pump: flow controller at lower limit', class Pump Warning Alarm, trigger "Pump5_Component_DBW_74" bit 12
   12538: 'Pump5: Component pump: max. filling level drip pan', class Pump Warning Alarm, trigger "Pump5_Component_DBW_74" bit 13
   12539: 'Pump5: Component pump:', class Pump Warning Alarm, trigger "Pump5_Component_DBW_74" bit 14
   12540: 'Pump5: Component pump:', class Pump Warning Alarm, trigger "Pump5_Component_DBW_74" bit 15
   12541: 'Pump5: Component pump:', class Pump Warning Alarm, trigger "Pump5_Component_DBW_74" bit 0
   12542: 'Pump5: Component pump:', class Pump Warning Alarm, trigger "Pump5_Component_DBW_74" bit 1
   12543: 'Pump5: Component pump:', class Pump Warning Alarm, trigger "Pump5_Component_DBW_74" bit 2
   12544: 'Pump5: Component pump:', class Pump Warning Alarm, trigger "Pump5_Component_DBW_74" bit 3
   12545: 'Pump5: Component pump:', class Pump Warning Alarm, trigger "Pump5_Component_DBW_74" bit 4
   12546: 'Pump5: Component pump:', class Pump Warning Alarm, trigger "Pump5_Component_DBW_74" bit 5
   12547: 'Pump5: Component pump:', class Pump Warning Alarm, trigger "Pump5_Component_DBW_74" bit 6
   12548: 'Pump5: Component pump:', class Pump Warning Alarm, trigger "Pump5_Component_DBW_74" bit 7
   12550: 'Pump5: Flow rate recording: measured value outside measuring range', class Pump Warning Alarm, trigger "Pump5_Flowrate_Record_DBW_114" bit 8
   12551: 'Pump5: Flow rate recording: warning, value exceeded', class Pump Warning Alarm, trigger "Pump5_Flowrate_Record_DBW_114" bit 9
   12552: 'Pump5: Flow rate recording: warning, value undershot', class Pump Warning Alarm, trigger "Pump5_Flowrate_Record_DBW_114" bit 10
   12553: 'Pump5: Flow rate recording: fault, value exceeded', class Pump Error Alarm, trigger "Pump5_Flowrate_Record_DBW_114" bit 11
   12554: 'Pump5: Flow rate recording: fault, value undershot', class Pump Error Alarm, trigger "Pump5_Flowrate_Record_DBW_114" bit 12
   12555: 'Pump5: Mixing ratio:', class Pump Warning Alarm, trigger "Pump5_Flowrate_Record_DBW_114" bit 0
   12556: 'Pump5: Mixing ratio: warning, value exceeded', class Pump Warning Alarm, trigger "Pump5_Flowrate_Record_DBW_114" bit 1
   12557: 'Pump5: Mixing ratio: warning, value undershot', class Pump Warning Alarm, trigger "Pump5_Flowrate_Record_DBW_114" bit 2
   12558: 'Pump5: Mixing ratio: fault, value exceeded', class Pump Error Alarm, trigger "Pump5_Flowrate_Record_DBW_114" bit 3
   12559: 'Pump5: Mixing ratio: fault, value undershot', class Pump Error Alarm, trigger "Pump5_Flowrate_Record_DBW_114" bit 4
   12560: 'Pump5: Pressure recording: measured value outside measuring range', class Pump Warning Alarm, trigger "Pump5_Pressure_Record_DBW_140" bit 8
   12561: 'Pump5: Pressure recording: warning, value exceeded', class Pump Warning Alarm, trigger "Pump5_Pressure_Record_DBW_140" bit 9
   12562: 'Pump5: Pressure recording: warning, value undershot', class Pump Warning Alarm, trigger "Pump5_Pressure_Record_DBW_140" bit 10
   12563: 'Pump5: Pressure recording: fault, value exceeded', class Pump Error Alarm, trigger "Pump5_Pressure_Record_DBW_140" bit 11
   12564: 'Pump5: Pressure recording: fault, value undershot', class Pump Error Alarm, trigger "Pump5_Pressure_Record_DBW_140" bit 12
   12565: 'Pump5: Temp. recording HP heat exch.: measured value outside measuring range', class Pump Warning Alarm, trigger "Pump5_Heatexchanger_DBW_218" bit 8
   12566: 'Pump5: Temp. recording HP heat exch.: warning, value exceeded', class Pump Warning Alarm, trigger "Pump5_Heatexchanger_DBW_218" bit 9
   12567: 'Pump5: Temp. recording HP heat exch.: warning, value undershot', class Pump Warning Alarm, trigger "Pump5_Heatexchanger_DBW_218" bit 10
   12568: 'Pump5: Temp. recording HP heat exch.: fault, value exceeded', class Pump Error Alarm, trigger "Pump5_Heatexchanger_DBW_218" bit 11
   12569: 'Pump5: Temp. recording HP heat exch.: fault, value undershot', class Pump Error Alarm, trigger "Pump5_Heatexchanger_DBW_218" bit 12
   12601: 'Pump6: FeedPump: motor protecting switch has tripped', class Pump Warning Alarm, trigger "Pump6_FeedPump_DBW_12" bit 8
   12602: 'Pump6: FeedPump: frequency converter fault', class Pump Warning Alarm, trigger "Pump6_FeedPump_DBW_12" bit 9
   12603: 'Pump6: FeedPump: max. filling level drip pan', class Pump Warning Alarm, trigger "Pump6_FeedPump_DBW_12" bit 10
   12604: 'Pump6: FeedPump: dry-run protection', class Pump Warning Alarm, trigger "Pump6_FeedPump_DBW_12" bit 11
   12605: 'Pump6: FeedPump: incorrect time entry for runtime or pause time', class Pump Warning Alarm, trigger "Pump6_FeedPump_DBW_12" bit 12
   12606: 'Pump6: FeedPump: temperature for switch-off not reached', class Pump Warning Alarm, trigger "Pump6_FeedPump_DBW_12" bit 13
   12607: 'Pump6: FeedPump: fan motor protecting switch', class Pump Warning Alarm, trigger "Pump6_FeedPump_DBW_12" bit 14
   12608: 'Pump6: FeedPump: filling level too low', class Pump Warning Alarm, trigger "Pump6_FeedPump_DBW_12" bit 15
   12609: 'Pump6: FeedPump:', class Pump Warning Alarm, trigger "Pump6_FeedPump_DBW_12" bit 0
   12610: 'Pump6: FeedPump: filling selected but no barrel present', class Pump Warning Alarm, trigger "Pump6_FeedPump_DBW_12" bit 1
   12611: 'Pump6: FeedPump: no barrel present', class Pump Warning Alarm, trigger "Pump6_FeedPump_DBW_12" bit 2
   12612: 'Pump6: FeedPump:', class Pump Warning Alarm, trigger "Pump6_FeedPump_DBW_12" bit 3
   12613: 'Pump6: EdgeFilter: motor protecting switch has tripped', class Pump Warning Alarm, trigger "Pump6_EdgeFilter_DBW_38" bit 8
   12614: 'Pump6: EdgeFilter: max. differential pressure', class Pump Warning Alarm, trigger "Pump6_EdgeFilter_DBW_38" bit 9
   12615: 'Pump6: EdgeFilter: incorrect time entry for runtime or pause time', class Pump Warning Alarm, trigger "Pump6_EdgeFilter_DBW_38" bit 10
   12616: 'Pump6: EdgeFilter:', class Pump Warning Alarm, trigger "Pump6_EdgeFilter_DBW_38" bit 11
   12617: 'Pump6: Component pump: admission pressure not present', class Pump Error Alarm, trigger "Pump6_Component_DBW_76" bit 8
   12618: 'Pump6: Component pump: motor protecting switch has tripped: Component pump', class Pump Error Alarm, trigger "Pump6_Component_DBW_76" bit 9
   12619: 'Pump6: Component pump: max. pressure', class Pump Error Alarm, trigger "Pump6_Component_DBW_76" bit 10
   12620: 'Pump6: Component pump: pressure after feedpump too low', class Pump Error Alarm, trigger "Pump6_Component_DBW_76" bit 11
   12621: 'Pump6: Component pump: frequency converter fault', class Pump Warning Alarm, trigger "Pump6_Component_DBW_76" bit 12
   12622: 'Pump6: Component pump: fan motor protecting switch', class Pump Warning Alarm, trigger "Pump6_Component_DBW_76" bit 13
   12623: 'Pump6: Component pump: min. tank filling level', class Pump Warning Alarm, trigger "Pump6_Component_DBW_76" bit 14
   12624: 'Pump6: Component pump: min. pressure not reached', class Pump Warning Alarm, trigger "Pump6_Component_DBW_76" bit 15
   12625: 'Pump6: Component pump: pre-alarm, nitrogen', class Pump Warning Alarm, trigger "Pump6_Component_DBW_76" bit 0
   12626: 'Pump6: Component pump: flow- tolerance +', class Pump Warning Alarm, trigger "Pump6_Component_DBW_76" bit 1
   12627: 'Pump6: Component pump: flow tolerance -', class Pump Warning Alarm, trigger "Pump6_Component_DBW_76" bit 2
   12628: 'Pump6: Component pump: Timeout at fast pressure build-up', class Pump Warning Alarm, trigger "Pump6_Component_DBW_76" bit 3
   12629: 'Pump6: Component pump: enable temperature not reached', class Pump Warning Alarm, trigger "Pump6_Component_DBW_76" bit 4
   12630: 'Pump6: Component pump: converter restart delay active', class Pump Warning Alarm, trigger "Pump6_Component_DBW_76" bit 5
   12631: 'Pump6: Component pump: alarm, nitrogen', class Pump Warning Alarm, trigger "Pump6_Component_DBW_76" bit 6
   12632: 'Pump6: Component pump: flow controller at limit', class Pump Warning Alarm, trigger "Pump6_Component_DBW_76" bit 7
   12633: 'Pump6: Component pump: component section was deselected', class Pump Warning Alarm, trigger "Pump6_Component_DBW_78" bit 8
   12634: 'Pump6: Component pump: deselected component section in interval', class Pump Warning Alarm, trigger "Pump6_Component_DBW_78" bit 9
   12635: 'Pump6: Component pump: fan motor protecting switch', class Pump Warning Alarm, trigger "Pump6_Component_DBW_78" bit 10
   12636: 'Pump6: Component pump: deselected component is required for entry', class Pump Warning Alarm, trigger "Pump6_Component_DBW_78" bit 11
   12637: 'Pump6: Component pump: flow controller at lower limit', class Pump Warning Alarm, trigger "Pump6_Component_DBW_78" bit 12
   12638: 'Pump6: Component pump: max. filling level drip pan', class Pump Warning Alarm, trigger "Pump6_Component_DBW_78" bit 13
   12639: 'Pump6: Component pump:', class Pump Warning Alarm, trigger "Pump6_Component_DBW_78" bit 14
   12640: 'Pump6: Component pump:', class Pump Warning Alarm, trigger "Pump6_Component_DBW_78" bit 15
   12641: 'Pump6: Component pump:', class Pump Warning Alarm, trigger "Pump6_Component_DBW_78" bit 0
   12642: 'Pump6: Component pump:', class Pump Warning Alarm, trigger "Pump6_Component_DBW_78" bit 1
   12643: 'Pump6: Component pump:', class Pump Warning Alarm, trigger "Pump6_Component_DBW_78" bit 2
   12644: 'Pump6: Component pump:', class Pump Warning Alarm, trigger "Pump6_Component_DBW_78" bit 3
   12645: 'Pump6: Component pump:', class Pump Warning Alarm, trigger "Pump6_Component_DBW_78" bit 4
   12646: 'Pump6: Component pump:', class Pump Warning Alarm, trigger "Pump6_Component_DBW_78" bit 5
   12647: 'Pump6: Component pump:', class Pump Warning Alarm, trigger "Pump6_Component_DBW_78" bit 6
   12648: 'Pump6: Component pump:', class Pump Warning Alarm, trigger "Pump6_Component_DBW_78" bit 7
   12650: 'Pump6: Flow rate recording: measured value outside measuring range', class Pump Warning Alarm, trigger "Pump6_Flowrate_Record_DBW_116" bit 8
   12651: 'Pump6: Flow rate recording: warning, value exceeded', class Pump Warning Alarm, trigger "Pump6_Flowrate_Record_DBW_116" bit 9
   12652: 'Pump6: Flow rate recording: warning, value undershot', class Pump Warning Alarm, trigger "Pump6_Flowrate_Record_DBW_116" bit 10
   12653: 'Pump6: Flow rate recording: fault, value exceeded', class Pump Error Alarm, trigger "Pump6_Flowrate_Record_DBW_116" bit 11
   12654: 'Pump6: Flow rate recording: fault, value undershot', class Pump Error Alarm, trigger "Pump6_Flowrate_Record_DBW_116" bit 12
   12655: 'Pump6: Mixing ratio:', class Pump Warning Alarm, trigger "Pump6_Flowrate_Record_DBW_116" bit 0
   12656: 'Pump6: Mixing ratio: warning, value exceeded', class Pump Warning Alarm, trigger "Pump6_Flowrate_Record_DBW_116" bit 1
   12657: 'Pump6: Mixing ratio: warning, value undershot', class Pump Warning Alarm, trigger "Pump6_Flowrate_Record_DBW_116" bit 2
   12658: 'Pump6: Mixing ratio: fault, value exceeded', class Pump Error Alarm, trigger "Pump6_Flowrate_Record_DBW_116" bit 3
   12659: 'Pump6: Mixing ratio: fault, value undershot', class Pump Error Alarm, trigger "Pump6_Flowrate_Record_DBW_116" bit 4
   12660: 'Pump6: Pressure recording: measured value outside measuring range', class Pump Warning Alarm, trigger "Pump6_Pressure_Record_DBW_142" bit 8
   12661: 'Pump6: Pressure recording: warning, value exceeded', class Pump Warning Alarm, trigger "Pump6_Pressure_Record_DBW_142" bit 9
